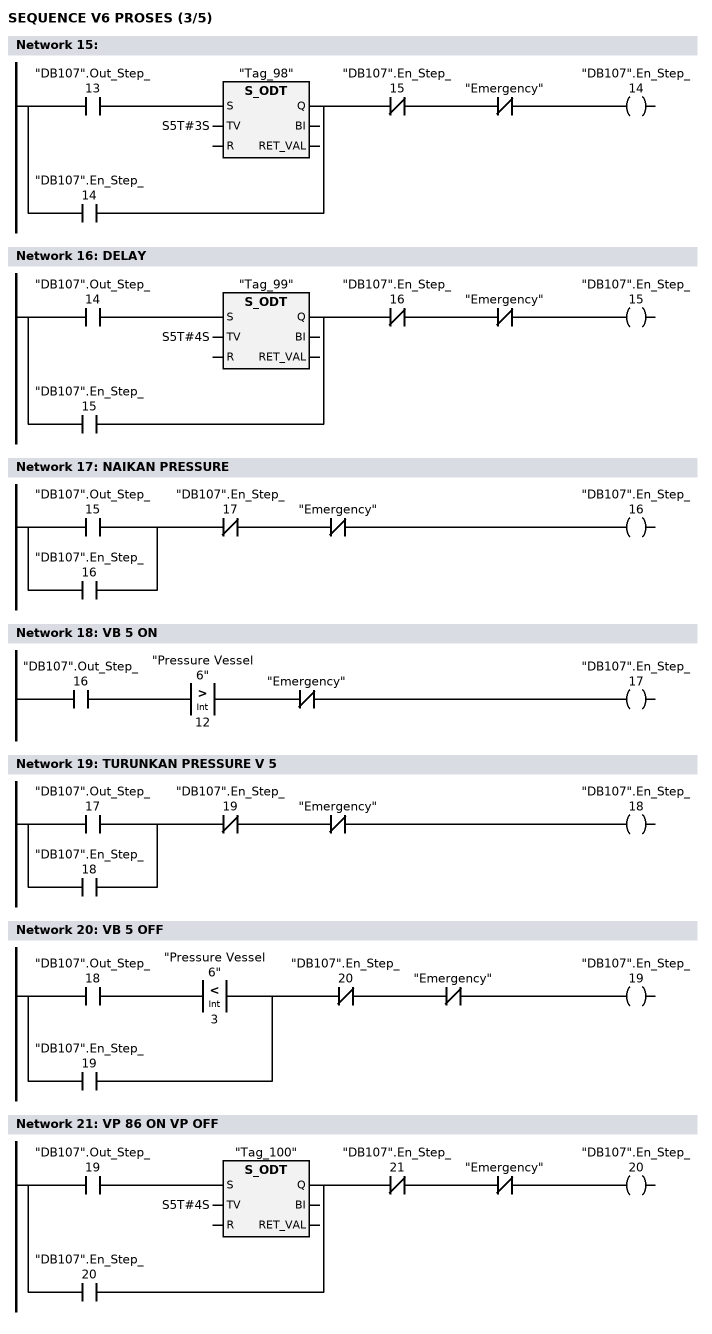
   RUNG wire#powerrail
      Contact( "DB107".Out_Step_13 )
      S_ODT(T_NO := "Tag_98", TV := S5T#3S, R :=, BI =>, RET_VAL =>)
      wire#w1
      I_Contact( "DB107".En_Step_15 )
      I_Contact( "Emergency" )
      Coil( "DB107".En_Step_14 )
   END_RUNG
   RUNG wire#powerrail
      Contact( "DB107".En_Step_14 )
   END_RUNG wire#w1
   // the same network as SCL:
   #_s5time1 := S_ODT(T_NO := "Tag_98", S := "DB107".Out_Step_13, TV := S5T#3S, Q => #_w1);
   "DB107".En_Step_14 := (#_w1 OR "DB107".En_Step_14) AND NOT "DB107".En_Step_15 AND NOT "Emergency";
END_REGION

REGION Network 16: DELAY
   RUNG wire#powerrail
      Contact( "DB107".Out_Step_14 )
      S_ODT(T_NO := "Tag_99", TV := S5T#4S, R :=, BI =>, RET_VAL =>)
      wire#w1
      I_Contact( "DB107".En_Step_16 )
      I_Contact( "Emergency" )
      Coil( "DB107".En_Step_15 )
   END_RUNG
   RUNG wire#powerrail
      Contact( "DB107".En_Step_15 )
   END_RUNG wire#w1
   // the same network as SCL:
   #_s5time1 := S_ODT(T_NO := "Tag_99", S := "DB107".Out_Step_14, TV := S5T#4S, Q => #_w1);
   "DB107".En_Step_15 := (#_w1 OR "DB107".En_Step_15) AND NOT "DB107".En_Step_16 AND NOT "Emergency";
END_REGION

REGION Network 17: NAIKAN PRESSURE
   RUNG wire#powerrail
      Contact( "DB107".Out_Step_15 )
      wire#w1
      I_Contact( "DB107".En_Step_17 )
      I_Contact( "Emergency" )
      Coil( "DB107".En_Step_16 )
   END_RUNG
   RUNG wire#powerrail
      Contact( "DB107".En_Step_16 )
   END_RUNG wire#w1
   // the same network as SCL:
   "DB107".En_Step_16 := ("DB107".Out_Step_15 OR "DB107".En_Step_16) AND NOT "DB107".En_Step_17 AND NOT "Emergency";
END_REGION

REGION Network 18: VB 5 ON
   RUNG wire#powerrail
      Contact( "DB107".Out_Step_16 )
      { S7_Templates := "SrcType := Int" } GT_Contact(in1 := "Pressure Vessel 6", in2 := 12)
      I_Contact( "Emergency" )
      Coil( "DB107".En_Step_17 )
   END_RUNG
   // the same network as SCL:
   "DB107".En_Step_17 := "DB107".Out_Step_16 AND ("Pressure Vessel 6" > 12) AND NOT "Emergency";
END_REGION

REGION Network 19: TURUNKAN PRESSURE V 5
   RUNG wire#powerrail
      Contact( "DB107".Out_Step_17 )
      wire#w1
      I_Contact( "DB107".En_Step_19 )
      I_Contact( "Emergency" )
      Coil( "DB107".En_Step_18 )
   END_RUNG
   RUNG wire#powerrail
      Contact( "DB107".En_Step_18 )
   END_RUNG wire#w1
   // the same network as SCL:
   "DB107".En_Step_18 := ("DB107".Out_Step_17 OR "DB107".En_Step_18) AND NOT "DB107".En_Step_19 AND NOT "Emergency";
END_REGION

REGION Network 20: VB 5 OFF
   RUNG wire#powerrail
      Contact( "DB107".Out_Step_18 )
      { S7_Templates := "SrcType := Int" } LT_Contact(in1 := "Pressure Vessel 6", in2 := 3)
      wire#w1
      I_Contact( "DB107".En_Step_20 )
      I_Contact( "Emergency" )
      Coil( "DB107".En_Step_19 )
   END_RUNG
   RUNG wire#powerrail
      Contact( "DB107".En_Step_19 )
   END_RUNG wire#w1
   // the same network as SCL:
   "DB107".En_Step_19 := (("DB107".Out_Step_18 AND ("Pressure Vessel 6" < 3)) OR "DB107".En_Step_19) AND NOT "DB107".En_Step_20 AND NOT "Emergency";
END_REGION

REGION Network 21: VP 86 ON VP OFF
   RUNG wire#powerrail
      Contact( "DB107".Out_Step_19 )
      S_ODT(T_NO := "Tag_100", TV := S5T#4S, R :=, BI =>, RET_VAL =>)
      wire#w1
      I_Contact( "DB107".En_Step_21 )
      I_Contact( "Emergency" )
      Coil( "DB107".En_Step_20 )
   END_RUNG
   RUNG wire#powerrail
      Contact( "DB107".En_Step_20 )
   END_RUNG wire#w1
   // the same network as SCL:
   #_s5time1 := S_ODT(T_NO := "Tag_100", S := "DB107".Out_Step_19, TV := S5T#4S, Q => #_w1);
   "DB107".En_Step_20 := (#_w1 OR "DB107".En_Step_20) AND NOT "DB107".En_Step_21 AND NOT "Emergency";
END_REGION

REGION Network 22: VP 86 OFF VP 87 ON
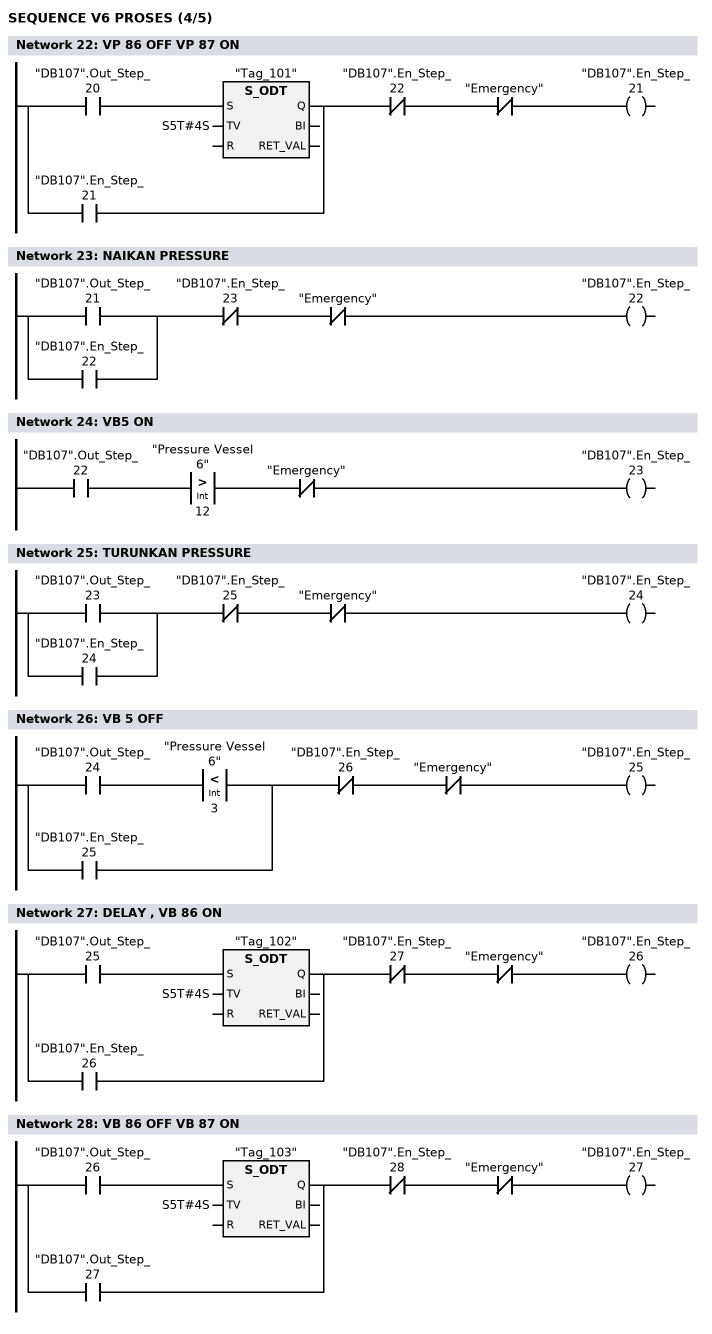
   RUNG wire#powerrail
      Contact( "DB107".Out_Step_20 )
      S_ODT(T_NO := "Tag_101", TV := S5T#4S, R :=, BI =>, RET_VAL =>)
      wire#w1
      I_Contact( "DB107".En_Step_22 )
      I_Contact( "Emergency" )
      Coil( "DB107".En_Step_21 )
   END_RUNG
   RUNG wire#powerrail
      Contact( "DB107".En_Step_21 )
   END_RUNG wire#w1
   // the same network as SCL:
   #_s5time1 := S_ODT(T_NO := "Tag_101", S := "DB107".Out_Step_20, TV := S5T#4S, Q => #_w1);
   "DB107".En_Step_21 := (#_w1 OR "DB107".En_Step_21) AND NOT "DB107".En_Step_22 AND NOT "Emergency";
END_REGION

REGION Network 23: NAIKAN PRESSURE
   RUNG wire#powerrail
      Contact( "DB107".Out_Step_21 )
      wire#w1
      I_Contact( "DB107".En_Step_23 )
      I_Contact( "Emergency" )
      Coil( "DB107".En_Step_22 )
   END_RUNG
   RUNG wire#powerrail
      Contact( "DB107".En_Step_22 )
   END_RUNG wire#w1
   // the same network as SCL:
   "DB107".En_Step_22 := ("DB107".Out_Step_21 OR "DB107".En_Step_22) AND NOT "DB107".En_Step_23 AND NOT "Emergency";
END_REGION

REGION Network 24: VB5 ON
   RUNG wire#powerrail
      Contact( "DB107".Out_Step_22 )
      { S7_Templates := "SrcType := Int" } GT_Contact(in1 := "Pressure Vessel 6", in2 := 12)
      I_Contact( "Emergency" )
      Coil( "DB107".En_Step_23 )
   END_RUNG
   // the same network as SCL:
   "DB107".En_Step_23 := "DB107".Out_Step_22 AND ("Pressure Vessel 6" > 12) AND NOT "Emergency";
END_REGION

REGION Network 25: TURUNKAN PRESSURE
   RUNG wire#powerrail
      Contact( "DB107".Out_Step_23 )
      wire#w1
      I_Contact( "DB107".En_Step_25 )
      I_Contact( "Emergency" )
      Coil( "DB107".En_Step_24 )
   END_RUNG
   RUNG wire#powerrail
      Contact( "DB107".En_Step_24 )
   END_RUNG wire#w1
   // the same network as SCL:
   "DB107".En_Step_24 := ("DB107".Out_Step_23 OR "DB107".En_Step_24) AND NOT "DB107".En_Step_25 AND NOT "Emergency";
END_REGION

REGION Network 26: VB 5 OFF
   RUNG wire#powerrail
      Contact( "DB107".Out_Step_24 )
      { S7_Templates := "SrcType := Int" } LT_Contact(in1 := "Pressure Vessel 6", in2 := 3)
      wire#w1
      I_Contact( "DB107".En_Step_26 )
      I_Contact( "Emergency" )
      Coil( "DB107".En_Step_25 )
   END_RUNG
   RUNG wire#powerrail
      Contact( "DB107".En_Step_25 )
   END_RUNG wire#w1
   // the same network as SCL:
   "DB107".En_Step_25 := (("DB107".Out_Step_24 AND ("Pressure Vessel 6" < 3)) OR "DB107".En_Step_25) AND NOT "DB107".En_Step_26 AND NOT "Emergency";
END_REGION

REGION Network 27: DELAY , VB 86 ON
   RUNG wire#powerrail
      Contact( "DB107".Out_Step_25 )
      S_ODT(T_NO := "Tag_102", TV := S5T#4S, R :=, BI =>, RET_VAL =>)
      wire#w1
      I_Contact( "DB107".En_Step_27 )
      I_Contact( "Emergency" )
      Coil( "DB107".En_Step_26 )
   END_RUNG
   RUNG wire#powerrail
      Contact( "DB107".En_Step_26 )
   END_RUNG wire#w1
   // the same network as SCL:
   #_s5time1 := S_ODT(T_NO := "Tag_102", S := "DB107".Out_Step_25, TV := S5T#4S, Q => #_w1);
   "DB107".En_Step_26 := (#_w1 OR "DB107".En_Step_26) AND NOT "DB107".En_Step_27 AND NOT "Emergency";
END_REGION

REGION Network 28: VB 86 OFF VB 87 ON
   RUNG wire#powerrail
      Contact( "DB107".Out_Step_26 )
      S_ODT(T_NO := "Tag_103", TV := S5T#4S, R :=, BI =>, RET_VAL =>)
      wire#w1
      I_Contact( "DB107".En_Step_28 )
      I_Contact( "Emergency" )
      Coil( "DB107".En_Step_27 )
   END_RUNG
   RUNG wire#powerrail
      Contact( "DB107".Out_Step_27 )
   END_RUNG wire#w1
   // the same network as SCL:
   #_s5time1 := S_ODT(T_NO := "Tag_103", S := "DB107".Out_Step_26, TV := S5T#4S, Q => #_w1);
   "DB107".En_Step_27 := (#_w1 OR "DB107".Out_Step_27) AND NOT "DB107".En_Step_28 AND NOT "Emergency";
END_REGION

REGION Network 29
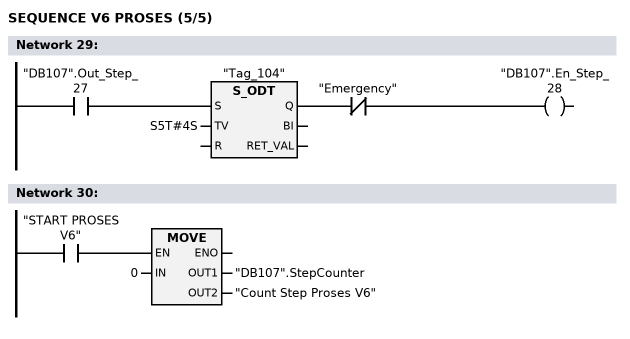
   RUNG wire#powerrail
      Contact( "DB107".Out_Step_27 )
      S_ODT(T_NO := "Tag_104", TV := S5T#4S, R :=, BI =>, RET_VAL =>)
      I_Contact( "Emergency" )
      Coil( "DB107".En_Step_28 )
   END_RUNG
   // the same network as SCL:
   #_s5time1 := S_ODT(T_NO := "Tag_104", S := "DB107".Out_Step_27, TV := S5T#4S, Q => #_w1);
   "DB107".En_Step_28 := #_w1 AND NOT "Emergency";
END_REGION

REGION Network 30
   RUNG wire#powerrail
      Contact( "START PROSES V6" )
      Move(in := 0, out1 => "DB107".StepCounter, out2 => "Count Step Proses V6")
   END_RUNG
   // the same network as SCL:
   IF "START PROSES V6" THEN
       "DB107".StepCounter := 0;
       "Count Step Proses V6" := 0;
   END_IF;
END_REGION
END_FUNCTION

FUNCTION "VESSEL 7 PROSES" : Void   // FC21, LAD
{ S7_Optimized_Access := 'TRUE' }
VERSION : 0.1
   VAR_TEMP   // added for the SCL form of the ladder/FBD networks
      _w1 : Bool;
      _w2 : Bool;
   END_VAR
BEGIN

REGION Network 1
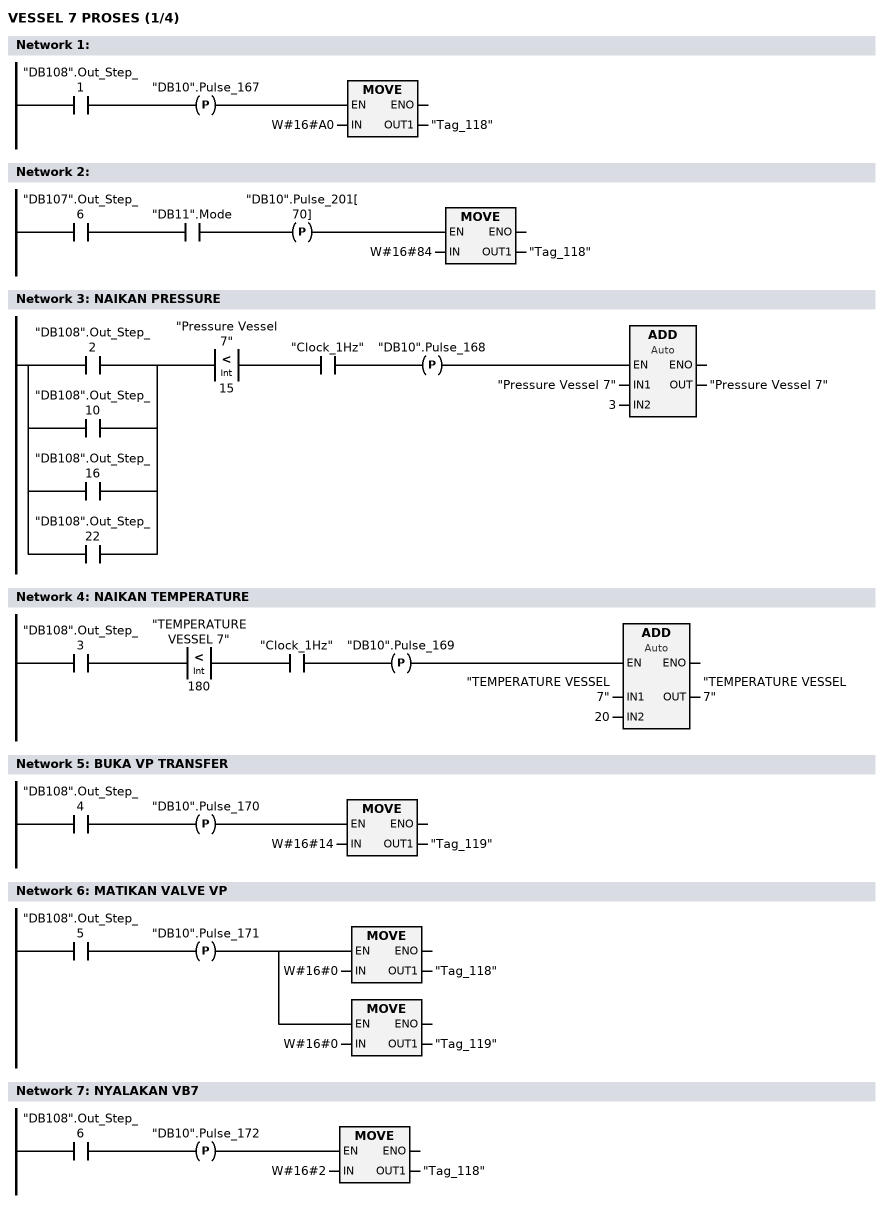
   RUNG wire#powerrail
      Contact( "DB108".Out_Step_1 )
      P_Trig( "DB10".Pulse_167 )
      Move(in := W#16#A0, out1 => "Tag_118")
   END_RUNG
   // the same network as SCL:
   #_w1 := "DB108".Out_Step_1 AND NOT "DB10".Pulse_167;   // rising edge
   "DB10".Pulse_167 := "DB108".Out_Step_1;
   IF #_w1 THEN "Tag_118" := W#16#A0; END_IF;
END_REGION

REGION Network 2
   RUNG wire#powerrail
      Contact( "DB107".Out_Step_6 )
      Contact( "DB11".Mode )
      P_Trig( "DB10".Pulse_201[70] )
      Move(in := W#16#84, out1 => "Tag_118")
   END_RUNG
   // the same network as SCL:
   #_w1 := "DB107".Out_Step_6 AND "DB11".Mode;
   #_w2 := #_w1 AND NOT "DB10".Pulse_201[70];   // rising edge
   "DB10".Pulse_201[70] := #_w1;
   IF #_w2 THEN "Tag_118" := W#16#84; END_IF;
END_REGION

REGION Network 3: NAIKAN PRESSURE
   RUNG wire#powerrail
      Contact( "DB108".Out_Step_2 )
      wire#w1
      { S7_Templates := "SrcType := Int" } LT_Contact(in1 := "Pressure Vessel 7", in2 := 15)
      Contact( "Clock_1Hz" )
      P_Trig( "DB10".Pulse_168 )
      Add(in1 := "Pressure Vessel 7", in2 := 3, out => "Pressure Vessel 7")
   END_RUNG
   RUNG wire#powerrail
      Contact( "DB108".Out_Step_10 )
   END_RUNG wire#w1
   RUNG wire#powerrail
      Contact( "DB108".Out_Step_16 )
   END_RUNG wire#w1
   RUNG wire#powerrail
      Contact( "DB108".Out_Step_22 )
   END_RUNG wire#w1
   // the same network as SCL:
   #_w1 := ("DB108".Out_Step_2 OR "DB108".Out_Step_10 OR "DB108".Out_Step_16 OR "DB108".Out_Step_22) AND ("Pressure Vessel 7" < 15) AND "Clock_1Hz";
   #_w2 := #_w1 AND NOT "DB10".Pulse_168;   // rising edge
   "DB10".Pulse_168 := #_w1;
   IF #_w2 THEN "Pressure Vessel 7" := "Pressure Vessel 7" + 3; END_IF;
END_REGION

REGION Network 4: NAIKAN TEMPERATURE
   RUNG wire#powerrail
      Contact( "DB108".Out_Step_3 )
      { S7_Templates := "SrcType := Int" } LT_Contact(in1 := "TEMPERATURE VESSEL 7", in2 := 180)
      Contact( "Clock_1Hz" )
      P_Trig( "DB10".Pulse_169 )
      Add(in1 := "TEMPERATURE VESSEL 7", in2 := 20, out => "TEMPERATURE VESSEL 7")
   END_RUNG
   // the same network as SCL:
   #_w1 := "DB108".Out_Step_3 AND ("TEMPERATURE VESSEL 7" < 180) AND "Clock_1Hz";
   #_w2 := #_w1 AND NOT "DB10".Pulse_169;   // rising edge
   "DB10".Pulse_169 := #_w1;
   IF #_w2 THEN "TEMPERATURE VESSEL 7" := "TEMPERATURE VESSEL 7" + 20; END_IF;
END_REGION

REGION Network 5: BUKA VP TRANSFER
   RUNG wire#powerrail
      Contact( "DB108".Out_Step_4 )
      P_Trig( "DB10".Pulse_170 )
      Move(in := W#16#14, out1 => "Tag_119")
   END_RUNG
   // the same network as SCL:
   #_w1 := "DB108".Out_Step_4 AND NOT "DB10".Pulse_170;   // rising edge
   "DB10".Pulse_170 := "DB108".Out_Step_4;
   IF #_w1 THEN "Tag_119" := W#16#14; END_IF;
END_REGION

REGION Network 6: MATIKAN VALVE VP
   RUNG wire#powerrail
      Contact( "DB108".Out_Step_5 )
      P_Trig( "DB10".Pulse_171 )
      wire#w1
      Move(in := W#16#0, out1 => "Tag_118")
   END_RUNG
   RUNG wire#w1
      Move(in := W#16#0, out1 => "Tag_119")
   END_RUNG
   // the same network as SCL:
   #_w1 := "DB108".Out_Step_5 AND NOT "DB10".Pulse_171;   // rising edge
   "DB10".Pulse_171 := "DB108".Out_Step_5;
   IF #_w1 THEN
       "Tag_118" := W#16#0;
       "Tag_119" := W#16#0;
   END_IF;
END_REGION

REGION Network 7: NYALAKAN VB7
   RUNG wire#powerrail
      Contact( "DB108".Out_Step_6 )
      P_Trig( "DB10".Pulse_172 )
      Move(in := W#16#2, out1 => "Tag_118")
   END_RUNG
   // the same network as SCL:
   #_w1 := "DB108".Out_Step_6 AND NOT "DB10".Pulse_172;   // rising edge
   "DB10".Pulse_172 := "DB108".Out_Step_6;
   IF #_w1 THEN "Tag_118" := W#16#2; END_IF;
END_REGION

REGION Network 8: TURUNKAN PRESSURE
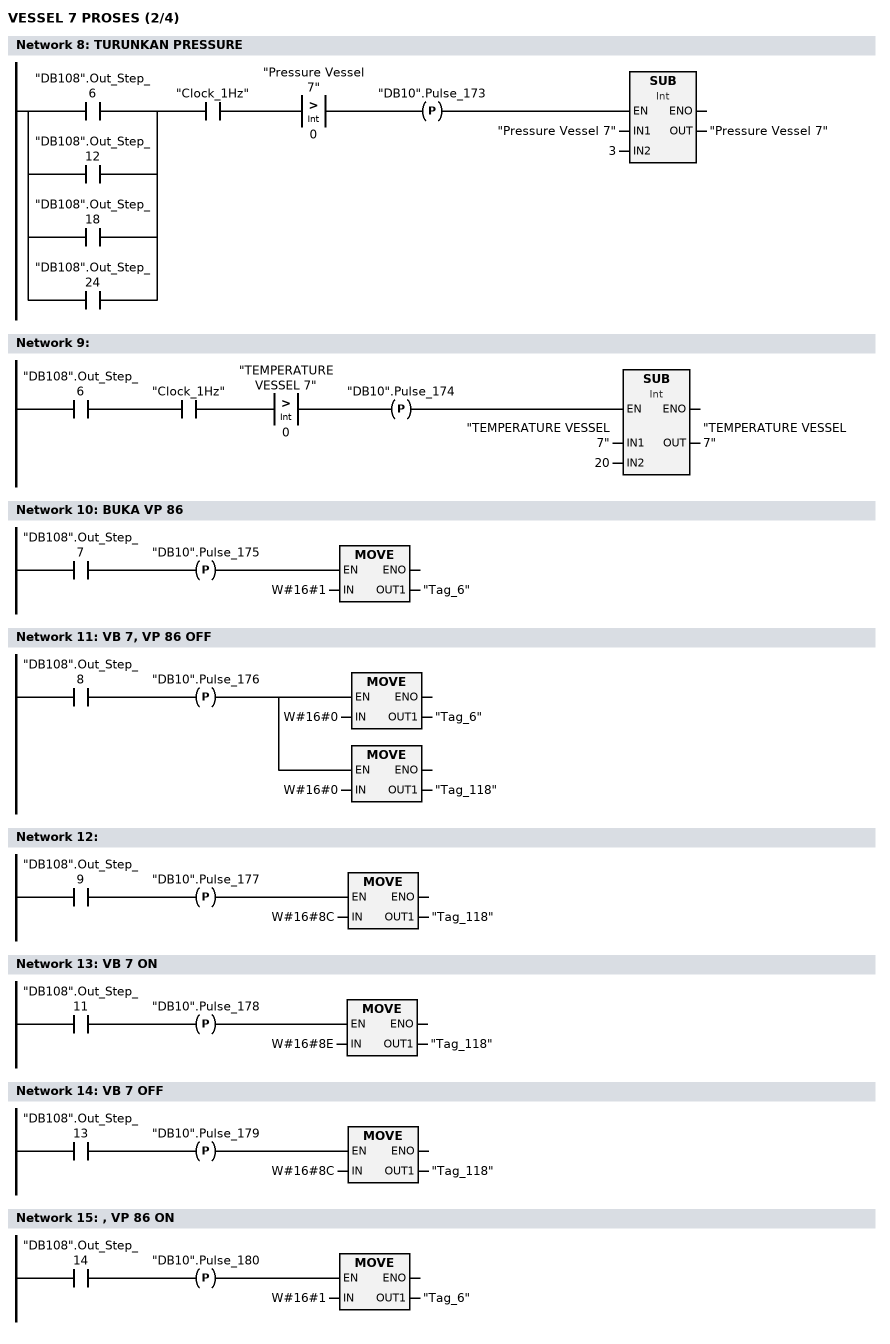
   RUNG wire#powerrail
      Contact( "DB108".Out_Step_6 )
      wire#w1
      Contact( "Clock_1Hz" )
      { S7_Templates := "SrcType := Int" } GT_Contact(in1 := "Pressure Vessel 7", in2 := 0)
      P_Trig( "DB10".Pulse_173 )
      { S7_Templates := "SrcType := Int" } Sub(in1 := "Pressure Vessel 7", in2 := 3, out => "Pressure Vessel 7")
   END_RUNG
   RUNG wire#powerrail
      Contact( "DB108".Out_Step_12 )
   END_RUNG wire#w1
   RUNG wire#powerrail
      Contact( "DB108".Out_Step_18 )
   END_RUNG wire#w1
   RUNG wire#powerrail
      Contact( "DB108".Out_Step_24 )
   END_RUNG wire#w1
   // the same network as SCL:
   #_w1 := ("DB108".Out_Step_6 OR "DB108".Out_Step_12 OR "DB108".Out_Step_18 OR "DB108".Out_Step_24) AND "Clock_1Hz" AND ("Pressure Vessel 7" > 0);
   #_w2 := #_w1 AND NOT "DB10".Pulse_173;   // rising edge
   "DB10".Pulse_173 := #_w1;
   IF #_w2 THEN "Pressure Vessel 7" := "Pressure Vessel 7" - 3; END_IF;
END_REGION

REGION Network 9
   RUNG wire#powerrail
      Contact( "DB108".Out_Step_6 )
      Contact( "Clock_1Hz" )
      { S7_Templates := "SrcType := Int" } GT_Contact(in1 := "TEMPERATURE VESSEL 7", in2 := 0)
      P_Trig( "DB10".Pulse_174 )
      { S7_Templates := "SrcType := Int" } Sub(in1 := "TEMPERATURE VESSEL 7", in2 := 20, out => "TEMPERATURE VESSEL 7")
   END_RUNG
   // the same network as SCL:
   #_w1 := "DB108".Out_Step_6 AND "Clock_1Hz" AND ("TEMPERATURE VESSEL 7" > 0);
   #_w2 := #_w1 AND NOT "DB10".Pulse_174;   // rising edge
   "DB10".Pulse_174 := #_w1;
   IF #_w2 THEN "TEMPERATURE VESSEL 7" := "TEMPERATURE VESSEL 7" - 20; END_IF;
END_REGION

REGION Network 10: BUKA VP 86
   RUNG wire#powerrail
      Contact( "DB108".Out_Step_7 )
      P_Trig( "DB10".Pulse_175 )
      Move(in := W#16#1, out1 => "Tag_6")
   END_RUNG
   // the same network as SCL:
   #_w1 := "DB108".Out_Step_7 AND NOT "DB10".Pulse_175;   // rising edge
   "DB10".Pulse_175 := "DB108".Out_Step_7;
   IF #_w1 THEN "Tag_6" := W#16#1; END_IF;
END_REGION

REGION Network 11: VB 7, VP 86 OFF
   RUNG wire#powerrail
      Contact( "DB108".Out_Step_8 )
      P_Trig( "DB10".Pulse_176 )
      wire#w1
      Move(in := W#16#0, out1 => "Tag_6")
   END_RUNG
   RUNG wire#w1
      Move(in := W#16#0, out1 => "Tag_118")
   END_RUNG
   // the same network as SCL:
   #_w1 := "DB108".Out_Step_8 AND NOT "DB10".Pulse_176;   // rising edge
   "DB10".Pulse_176 := "DB108".Out_Step_8;
   IF #_w1 THEN
       "Tag_6" := W#16#0;
       "Tag_118" := W#16#0;
   END_IF;
END_REGION

REGION Network 12
   RUNG wire#powerrail
      Contact( "DB108".Out_Step_9 )
      P_Trig( "DB10".Pulse_177 )
      Move(in := W#16#8C, out1 => "Tag_118")
   END_RUNG
   // the same network as SCL:
   #_w1 := "DB108".Out_Step_9 AND NOT "DB10".Pulse_177;   // rising edge
   "DB10".Pulse_177 := "DB108".Out_Step_9;
   IF #_w1 THEN "Tag_118" := W#16#8C; END_IF;
END_REGION

REGION Network 13: VB 7 ON
   RUNG wire#powerrail
      Contact( "DB108".Out_Step_11 )
      P_Trig( "DB10".Pulse_178 )
      Move(in := W#16#8E, out1 => "Tag_118")
   END_RUNG
   // the same network as SCL:
   #_w1 := "DB108".Out_Step_11 AND NOT "DB10".Pulse_178;   // rising edge
   "DB10".Pulse_178 := "DB108".Out_Step_11;
   IF #_w1 THEN "Tag_118" := W#16#8E; END_IF;
END_REGION

REGION Network 14: VB 7 OFF
   RUNG wire#powerrail
      Contact( "DB108".Out_Step_13 )
      P_Trig( "DB10".Pulse_179 )
      Move(in := W#16#8C, out1 => "Tag_118")
   END_RUNG
   // the same network as SCL:
   #_w1 := "DB108".Out_Step_13 AND NOT "DB10".Pulse_179;   // rising edge
   "DB10".Pulse_179 := "DB108".Out_Step_13;
   IF #_w1 THEN "Tag_118" := W#16#8C; END_IF;
END_REGION

REGION Network 15: , VP 86 ON
   RUNG wire#powerrail
      Contact( "DB108".Out_Step_14 )
      P_Trig( "DB10".Pulse_180 )
      Move(in := W#16#1, out1 => "Tag_6")
   END_RUNG
   // the same network as SCL:
   #_w1 := "DB108".Out_Step_14 AND NOT "DB10".Pulse_180;   // rising edge
   "DB10".Pulse_180 := "DB108".Out_Step_14;
   IF #_w1 THEN "Tag_6" := W#16#1; END_IF;
END_REGION

REGION Network 16: VP 86 OFF
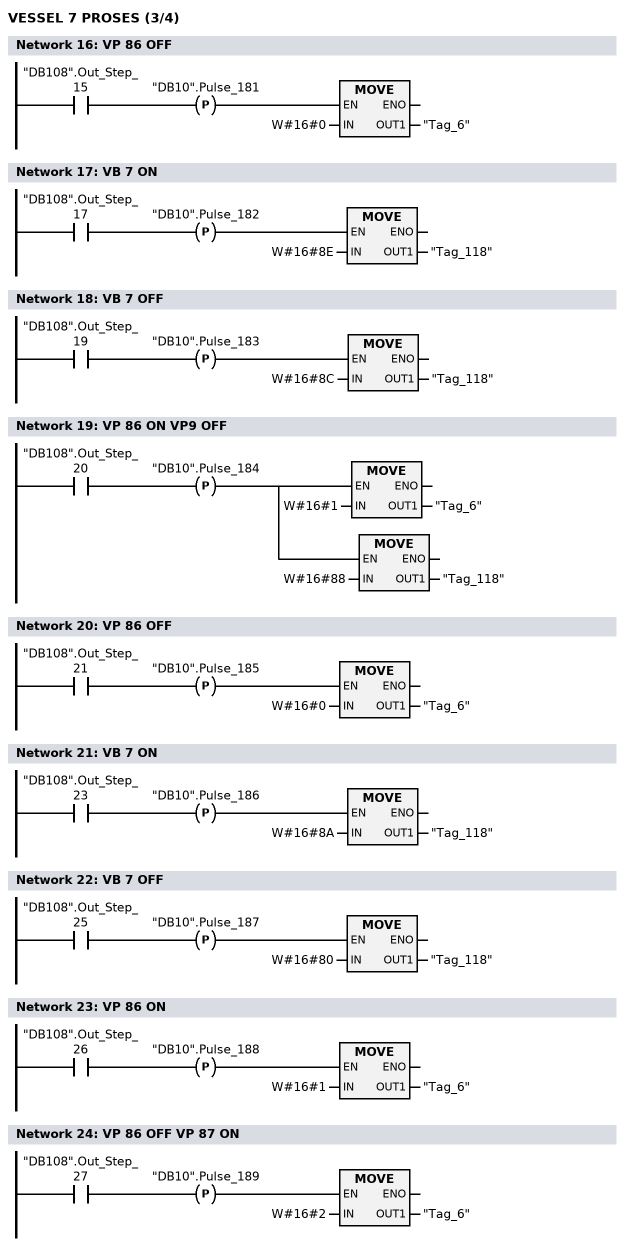
   RUNG wire#powerrail
      Contact( "DB108".Out_Step_15 )
      P_Trig( "DB10".Pulse_181 )
      Move(in := W#16#0, out1 => "Tag_6")
   END_RUNG
   // the same network as SCL:
   #_w1 := "DB108".Out_Step_15 AND NOT "DB10".Pulse_181;   // rising edge
   "DB10".Pulse_181 := "DB108".Out_Step_15;
   IF #_w1 THEN "Tag_6" := W#16#0; END_IF;
END_REGION

REGION Network 17: VB 7 ON
   RUNG wire#powerrail
      Contact( "DB108".Out_Step_17 )
      P_Trig( "DB10".Pulse_182 )
      Move(in := W#16#8E, out1 => "Tag_118")
   END_RUNG
   // the same network as SCL:
   #_w1 := "DB108".Out_Step_17 AND NOT "DB10".Pulse_182;   // rising edge
   "DB10".Pulse_182 := "DB108".Out_Step_17;
   IF #_w1 THEN "Tag_118" := W#16#8E; END_IF;
END_REGION

REGION Network 18: VB 7 OFF
   RUNG wire#powerrail
      Contact( "DB108".Out_Step_19 )
      P_Trig( "DB10".Pulse_183 )
      Move(in := W#16#8C, out1 => "Tag_118")
   END_RUNG
   // the same network as SCL:
   #_w1 := "DB108".Out_Step_19 AND NOT "DB10".Pulse_183;   // rising edge
   "DB10".Pulse_183 := "DB108".Out_Step_19;
   IF #_w1 THEN "Tag_118" := W#16#8C; END_IF;
END_REGION

REGION Network 19: VP 86 ON VP9 OFF
   RUNG wire#powerrail
      Contact( "DB108".Out_Step_20 )
      P_Trig( "DB10".Pulse_184 )
      wire#w1
      Move(in := W#16#1, out1 => "Tag_6")
   END_RUNG
   RUNG wire#w1
      Move(in := W#16#88, out1 => "Tag_118")
   END_RUNG
   // the same network as SCL:
   #_w1 := "DB108".Out_Step_20 AND NOT "DB10".Pulse_184;   // rising edge
   "DB10".Pulse_184 := "DB108".Out_Step_20;
   IF #_w1 THEN
       "Tag_6" := W#16#1;
       "Tag_118" := W#16#88;
   END_IF;
END_REGION

REGION Network 20: VP 86 OFF
   RUNG wire#powerrail
      Contact( "DB108".Out_Step_21 )
      P_Trig( "DB10".Pulse_185 )
      Move(in := W#16#0, out1 => "Tag_6")
   END_RUNG
   // the same network as SCL:
   #_w1 := "DB108".Out_Step_21 AND NOT "DB10".Pulse_185;   // rising edge
   "DB10".Pulse_185 := "DB108".Out_Step_21;
   IF #_w1 THEN "Tag_6" := W#16#0; END_IF;
END_REGION

REGION Network 21: VB 7 ON
   RUNG wire#powerrail
      Contact( "DB108".Out_Step_23 )
      P_Trig( "DB10".Pulse_186 )
      Move(in := W#16#8A, out1 => "Tag_118")
   END_RUNG
   // the same network as SCL:
   #_w1 := "DB108".Out_Step_23 AND NOT "DB10".Pulse_186;   // rising edge
   "DB10".Pulse_186 := "DB108".Out_Step_23;
   IF #_w1 THEN "Tag_118" := W#16#8A; END_IF;
END_REGION

REGION Network 22: VB 7 OFF
   RUNG wire#powerrail
      Contact( "DB108".Out_Step_25 )
      P_Trig( "DB10".Pulse_187 )
      Move(in := W#16#80, out1 => "Tag_118")
   END_RUNG
   // the same network as SCL:
   #_w1 := "DB108".Out_Step_25 AND NOT "DB10".Pulse_187;   // rising edge
   "DB10".Pulse_187 := "DB108".Out_Step_25;
   IF #_w1 THEN "Tag_118" := W#16#80; END_IF;
END_REGION

REGION Network 23: VP 86 ON
   RUNG wire#powerrail
      Contact( "DB108".Out_Step_26 )
      P_Trig( "DB10".Pulse_188 )
      Move(in := W#16#1, out1 => "Tag_6")
   END_RUNG
   // the same network as SCL:
   #_w1 := "DB108".Out_Step_26 AND NOT "DB10".Pulse_188;   // rising edge
   "DB10".Pulse_188 := "DB108".Out_Step_26;
   IF #_w1 THEN "Tag_6" := W#16#1; END_IF;
END_REGION

REGION Network 24: VP 86 OFF VP 87 ON
   RUNG wire#powerrail
      Contact( "DB108".Out_Step_27 )
      P_Trig( "DB10".Pulse_189 )
      Move(in := W#16#2, out1 => "Tag_6")
   END_RUNG
   // the same network as SCL:
   #_w1 := "DB108".Out_Step_27 AND NOT "DB10".Pulse_189;   // rising edge
   "DB10".Pulse_189 := "DB108".Out_Step_27;
   IF #_w1 THEN "Tag_6" := W#16#2; END_IF;
END_REGION

REGION Network 25: VP 87 OFF
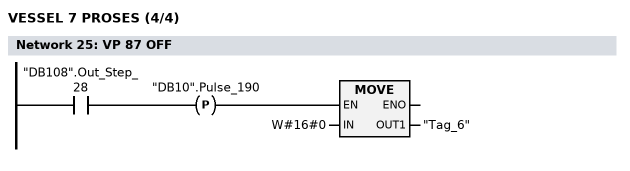
   RUNG wire#powerrail
      Contact( "DB108".Out_Step_28 )
      P_Trig( "DB10".Pulse_190 )
      Move(in := W#16#0, out1 => "Tag_6")
   END_RUNG
   // the same network as SCL:
   #_w1 := "DB108".Out_Step_28 AND NOT "DB10".Pulse_190;   // rising edge
   "DB10".Pulse_190 := "DB108".Out_Step_28;
   IF #_w1 THEN "Tag_6" := W#16#0; END_IF;
END_REGION
END_FUNCTION

FUNCTION "SEQUENCE V7 PROSES" : Void   // FC22, LAD
{ S7_Optimized_Access := 'TRUE' }
VERSION : 0.1
   VAR_TEMP   // added for the SCL form of the ladder/FBD networks
      _w1 : Bool;
      _w2 : Bool;
      _s5time1 : S5Time;
      _w3 : Bool;
   END_VAR
BEGIN

REGION Network 1: START PROSES
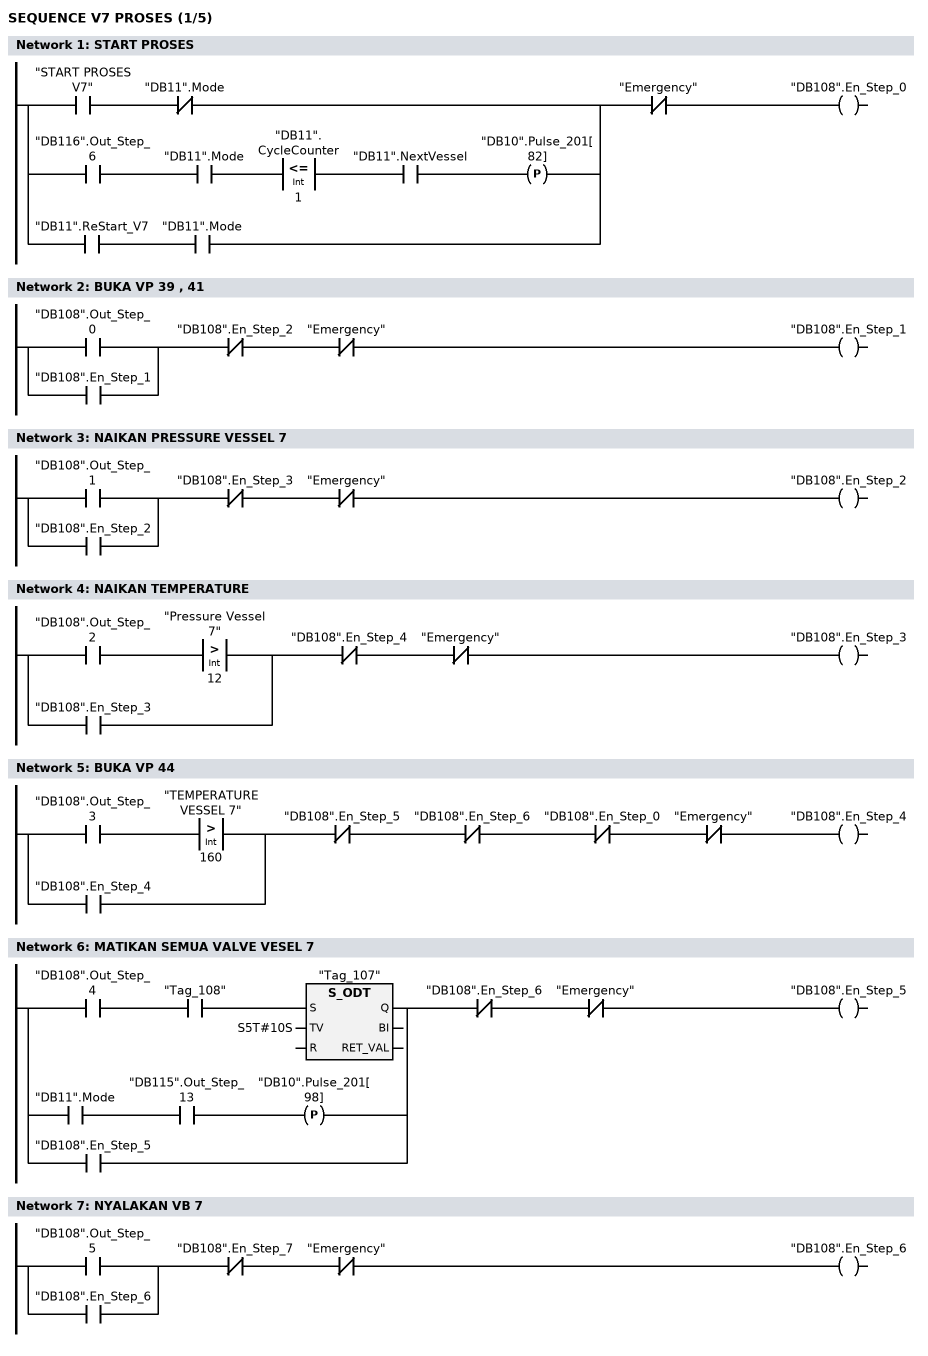
   RUNG wire#powerrail
      Contact( "START PROSES V7" )
      I_Contact( "DB11".Mode )
      wire#w1
      I_Contact( "Emergency" )
      Coil( "DB108".En_Step_0 )
   END_RUNG
   RUNG wire#powerrail
      Contact( "DB116".Out_Step_6 )
      Contact( "DB11".Mode )
      { S7_Templates := "SrcType := Int" } LE_Contact(in1 := "DB11".CycleCounter, in2 := 1)
      Contact( "DB11".NextVessel )
      P_Trig( "DB10".Pulse_201[82] )
   END_RUNG wire#w1
   RUNG wire#powerrail
      Contact( "DB11".ReStart_V7 )
      Contact( "DB11".Mode )
   END_RUNG wire#w1
   // the same network as SCL:
   #_w1 := "DB116".Out_Step_6 AND "DB11".Mode AND ("DB11".CycleCounter <= 1) AND "DB11".NextVessel;
   #_w2 := #_w1 AND NOT "DB10".Pulse_201[82];   // rising edge
   "DB10".Pulse_201[82] := #_w1;
   "DB108".En_Step_0 := (("START PROSES V7" AND NOT "DB11".Mode) OR #_w2 OR ("DB11".ReStart_V7 AND "DB11".Mode)) AND NOT "Emergency";
END_REGION

REGION Network 2: BUKA VP 39 , 41
   RUNG wire#powerrail
      Contact( "DB108".Out_Step_0 )
      wire#w1
      I_Contact( "DB108".En_Step_2 )
      I_Contact( "Emergency" )
      Coil( "DB108".En_Step_1 )
   END_RUNG
   RUNG wire#powerrail
      Contact( "DB108".En_Step_1 )
   END_RUNG wire#w1
   // the same network as SCL:
   "DB108".En_Step_1 := ("DB108".Out_Step_0 OR "DB108".En_Step_1) AND NOT "DB108".En_Step_2 AND NOT "Emergency";
END_REGION

REGION Network 3: NAIKAN PRESSURE VESSEL 7
   RUNG wire#powerrail
      Contact( "DB108".Out_Step_1 )
      wire#w1
      I_Contact( "DB108".En_Step_3 )
      I_Contact( "Emergency" )
      Coil( "DB108".En_Step_2 )
   END_RUNG
   RUNG wire#powerrail
      Contact( "DB108".En_Step_2 )
   END_RUNG wire#w1
   // the same network as SCL:
   "DB108".En_Step_2 := ("DB108".Out_Step_1 OR "DB108".En_Step_2) AND NOT "DB108".En_Step_3 AND NOT "Emergency";
END_REGION

REGION Network 4: NAIKAN TEMPERATURE
   RUNG wire#powerrail
      Contact( "DB108".Out_Step_2 )
      { S7_Templates := "SrcType := Int" } GT_Contact(in1 := "Pressure Vessel 7", in2 := 12)
      wire#w1
      I_Contact( "DB108".En_Step_4 )
      I_Contact( "Emergency" )
      Coil( "DB108".En_Step_3 )
   END_RUNG
   RUNG wire#powerrail
      Contact( "DB108".En_Step_3 )
   END_RUNG wire#w1
   // the same network as SCL:
   "DB108".En_Step_3 := (("DB108".Out_Step_2 AND ("Pressure Vessel 7" > 12)) OR "DB108".En_Step_3) AND NOT "DB108".En_Step_4 AND NOT "Emergency";
END_REGION

REGION Network 5: BUKA VP 44
   RUNG wire#powerrail
      Contact( "DB108".Out_Step_3 )
      { S7_Templates := "SrcType := Int" } GT_Contact(in1 := "TEMPERATURE VESSEL 7", in2 := 160)
      wire#w1
      I_Contact( "DB108".En_Step_5 )
      I_Contact( "DB108".En_Step_6 )
      I_Contact( "DB108".En_Step_0 )
      I_Contact( "Emergency" )
      Coil( "DB108".En_Step_4 )
   END_RUNG
   RUNG wire#powerrail
      Contact( "DB108".En_Step_4 )
   END_RUNG wire#w1
   // the same network as SCL:
   "DB108".En_Step_4 := (("DB108".Out_Step_3 AND ("TEMPERATURE VESSEL 7" > 160)) OR "DB108".En_Step_4) AND NOT "DB108".En_Step_5 AND NOT "DB108".En_Step_6 AND NOT "DB108".En_Step_0 AND NOT "Emergency";
END_REGION

REGION Network 6: MATIKAN SEMUA VALVE VESEL 7
   RUNG wire#powerrail
      Contact( "DB108".Out_Step_4 )
      Contact( "Tag_108" )
      S_ODT(T_NO := "Tag_107", TV := S5T#10S, R :=, BI =>, RET_VAL =>)
      wire#w1
      I_Contact( "DB108".En_Step_6 )
      I_Contact( "Emergency" )
      Coil( "DB108".En_Step_5 )
   END_RUNG
   RUNG wire#powerrail
      Contact( "DB11".Mode )
      Contact( "DB115".Out_Step_13 )
      P_Trig( "DB10".Pulse_201[98] )
   END_RUNG wire#w1
   RUNG wire#powerrail
      Contact( "DB108".En_Step_5 )
   END_RUNG wire#w1
   // the same network as SCL:
   #_s5time1 := S_ODT(T_NO := "Tag_107", S := "DB108".Out_Step_4 AND "Tag_108", TV := S5T#10S, Q => #_w1);
   #_w2 := "DB11".Mode AND "DB115".Out_Step_13;
   #_w3 := #_w2 AND NOT "DB10".Pulse_201[98];   // rising edge
   "DB10".Pulse_201[98] := #_w2;
   "DB108".En_Step_5 := (#_w1 OR #_w3 OR "DB108".En_Step_5) AND NOT "DB108".En_Step_6 AND NOT "Emergency";
END_REGION

REGION Network 7: NYALAKAN VB 7
   RUNG wire#powerrail
      Contact( "DB108".Out_Step_5 )
      wire#w1
      I_Contact( "DB108".En_Step_7 )
      I_Contact( "Emergency" )
      Coil( "DB108".En_Step_6 )
   END_RUNG
   RUNG wire#powerrail
      Contact( "DB108".En_Step_6 )
   END_RUNG wire#w1
   // the same network as SCL:
   "DB108".En_Step_6 := ("DB108".Out_Step_5 OR "DB108".En_Step_6) AND NOT "DB108".En_Step_7 AND NOT "Emergency";
END_REGION

REGION Network 8